(* Logix 5000 project; controller PLC_MCC1300_75F1 vendor 1 type 14 code 166 rev 32.11; software revision 32.04; part 51 of 83 *)
(* tags used below, declared in another part *)
   GP_ScadaPlate : GP_ScadaPlate;
   M310B : MAC_Conveyor;
   M310B_ALM : MAC_Conveyor_ALM;
   M310B_Data : UDT_Convoy_SL;
   M310B_HMR : MAC_Conveyor_HMR;
   M310B_SpaceConv_Utilities : SpaceConv_Utilities;
   M310Popup : MAC_Popup_ZC[2];
   M310Popup_ALM : MAC_Popup_ZC_ALM[2];
   M310Popup_HMR : MAC_Popup_ZC_HMR[2];
   M310Popup_HMW : MAC_Popup_ZC_HMW[2];
   TMP_dHalfConveyorLength : DINT;
   xAlwaysOFF : BOOL;
   xAlwaysON : BOOL;
   Z300_Conveyor : UDT_StandConv[29];
   Z300_LineTracking : UDT_LINE_TRACKING;
   Z301 : MAC_Zone_ML;
   Z401_HMI_rgtPlateScada_Internal : HMI_LiteData[5,2,7];
(* MainProgram, continued *)

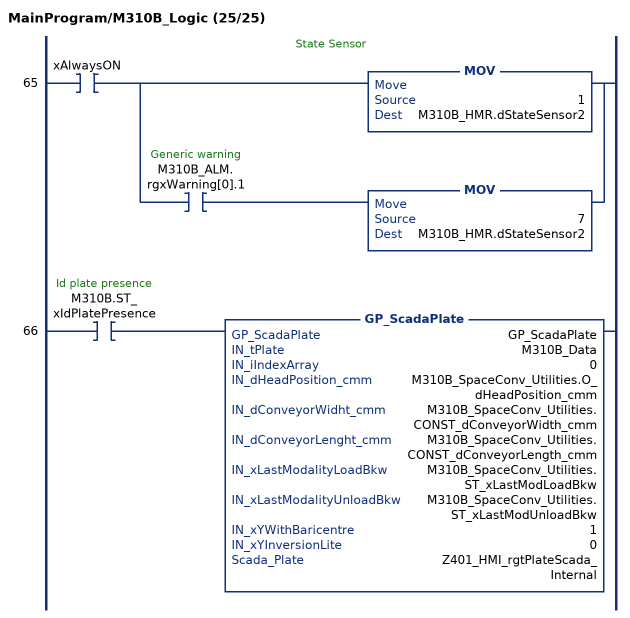
   [picture p787: MainProgram/M310B_Logic rungs 65-66]
   // State Sensor
   65: XIC(xAlwaysON)[MOV(1,M310B_HMR.dStateSensor2) ,XIC(M310B_ALM.rgxWarning[0].1) MOV(7,M310B_HMR.dStateSensor2) ];
   66: XIC(M310B.ST_xIdPlatePresence)GP_ScadaPlate(GP_ScadaPlate,M310B_Data,0,M310B_SpaceConv_Utilities.O_dHeadPosition_cmm,M310B_SpaceConv_Utilities.CONST_dConveyorWidth_cmm,M310B_SpaceConv_Utilities.CONST_dConveyorLength_cmm,M310B_SpaceConv_Utilities.ST_xLastModLoadBkw,M310B_SpaceConv_Utilities.ST_xLastModUnloadBkw,1,0,Z401_HMI_rgtPlateScada_Internal);
END_ROUTINE

ROUTINE M310Popup0_Faults   (* ladder *)
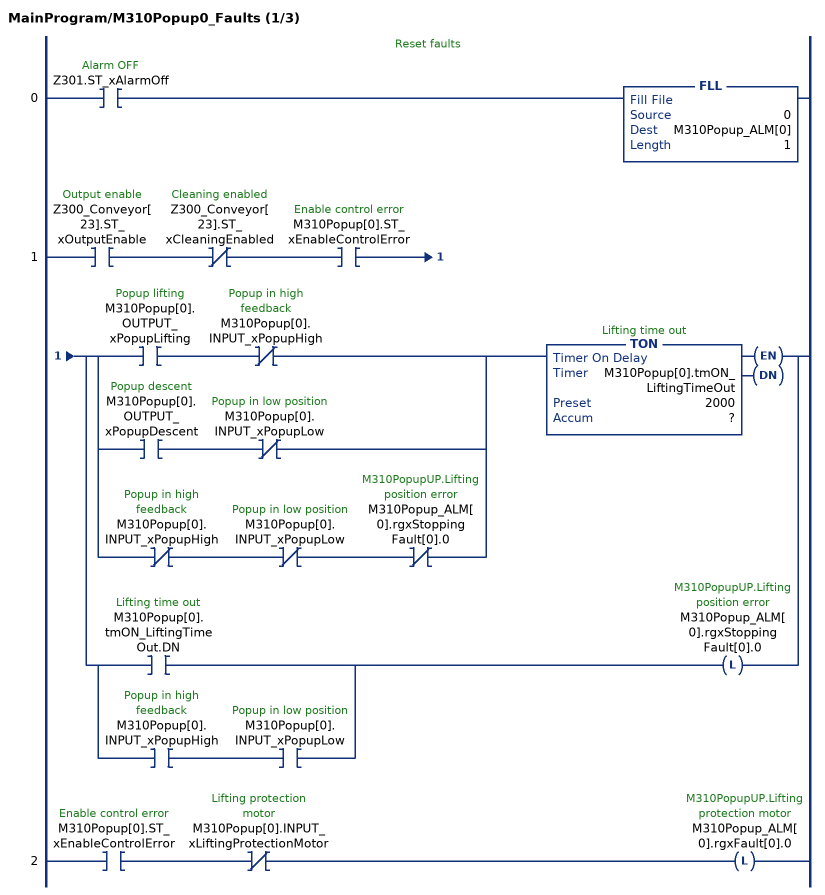
   // Reset faults
   0: XIC(Z301.ST_xAlarmOff)FLL(0,M310Popup_ALM[0],1);
   1: XIC(Z300_Conveyor[23].ST_xOutputEnable)XIO(Z300_Conveyor[23].ST_xCleaningEnabled)XIC(M310Popup[0].ST_xEnableControlError)[[XIC(M310Popup[0].OUTPUT_xPopupLifting) XIO(M310Popup[0].INPUT_xPopupHigh) ,XIC(M310Popup[0].OUTPUT_xPopupDescent) XIO(M310Popup[0].INPUT_xPopupLow) ,XIO(M310Popup[0].INPUT_xPopupHigh) XIO(M310Popup[0].INPUT_xPopupLow) XIO(M310Popup_ALM[0].rgxStoppingFault[0].0) ] TON(M310Popup[0].tmON_LiftingTimeOut,?,?) ,[XIC(M310Popup[0].tmON_LiftingTimeOut.DN) ,XIC(M310Popup[0].INPUT_xPopupHigh) XIC(M310Popup[0].INPUT_xPopupLow) ] OTL(M310Popup_ALM[0].rgxStoppingFault[0].0) ];
   2: XIC(M310Popup[0].ST_xEnableControlError)XIO(M310Popup[0].INPUT_xLiftingProtectionMotor)OTL(M310Popup_ALM[0].rgxFault[0].0);
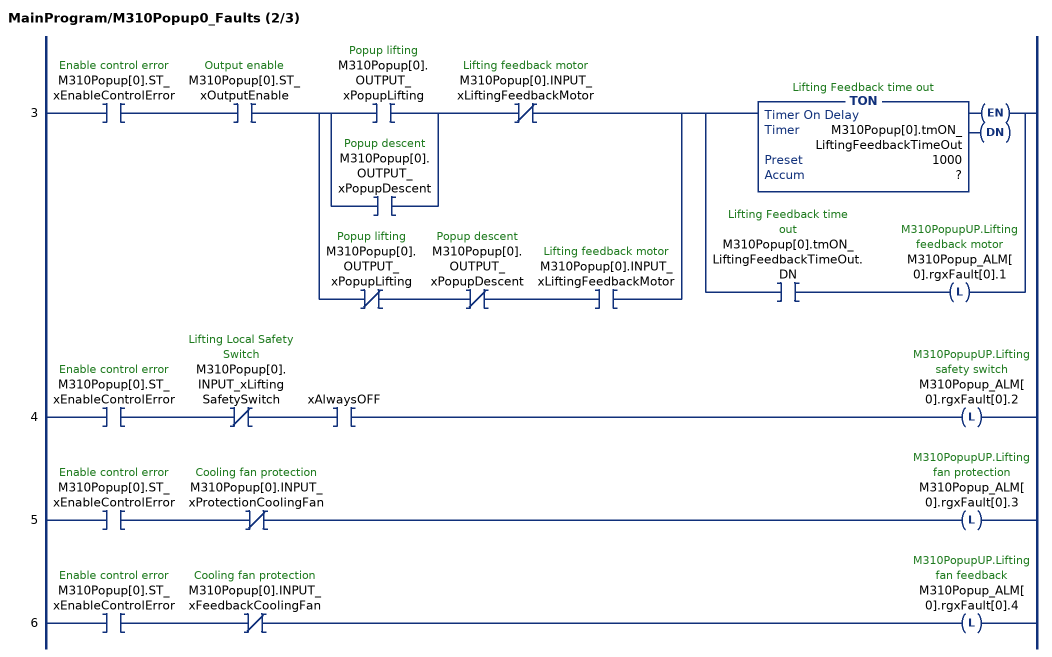
   3: XIC(M310Popup[0].ST_xEnableControlError)XIC(M310Popup[0].ST_xOutputEnable)[[XIC(M310Popup[0].OUTPUT_xPopupLifting) ,XIC(M310Popup[0].OUTPUT_xPopupDescent) ] XIO(M310Popup[0].INPUT_xLiftingFeedbackMotor) ,XIO(M310Popup[0].OUTPUT_xPopupLifting) XIO(M310Popup[0].OUTPUT_xPopupDescent) XIC(M310Popup[0].INPUT_xLiftingFeedbackMotor) ][TON(M310Popup[0].tmON_LiftingFeedbackTimeOut,?,?) ,XIC(M310Popup[0].tmON_LiftingFeedbackTimeOut.DN) OTL(M310Popup_ALM[0].rgxFault[0].1) ];
   4: XIC(M310Popup[0].ST_xEnableControlError)XIO(M310Popup[0].INPUT_xLiftingSafetySwitch)XIC(xAlwaysOFF)OTL(M310Popup_ALM[0].rgxFault[0].2);
   5: XIC(M310Popup[0].ST_xEnableControlError)XIO(M310Popup[0].INPUT_xProtectionCoolingFan)OTL(M310Popup_ALM[0].rgxFault[0].3);
   6: XIC(M310Popup[0].ST_xEnableControlError)XIO(M310Popup[0].INPUT_xFeedbackCoolingFan)OTL(M310Popup_ALM[0].rgxFault[0].4);
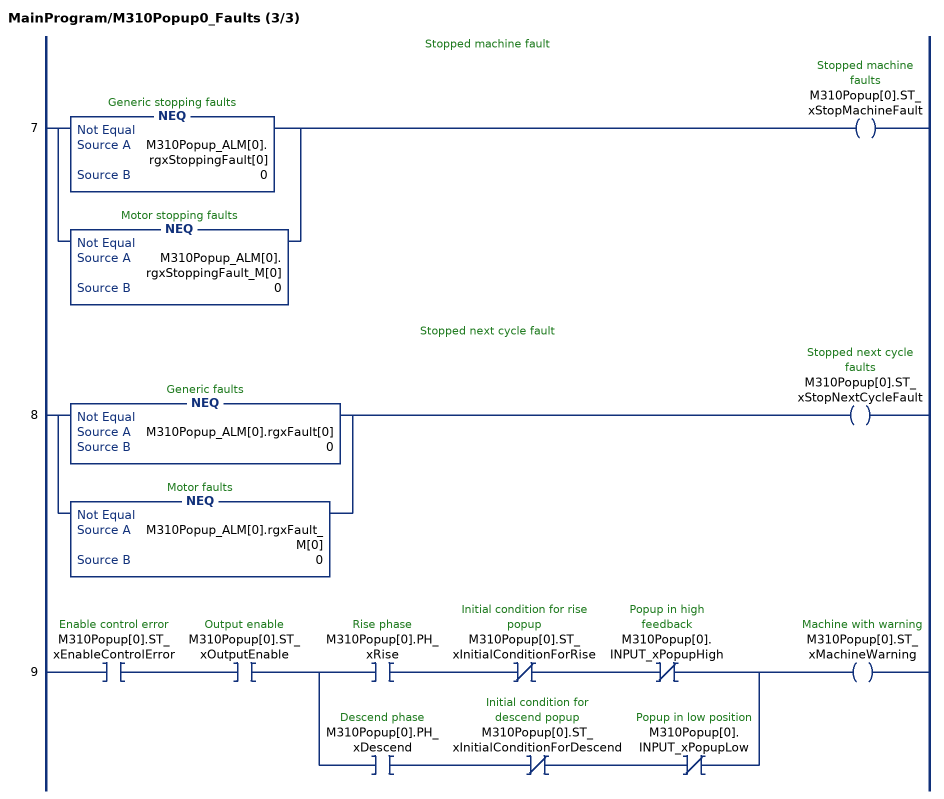
   // Stopped machine fault
   7: [NEQ(M310Popup_ALM[0].rgxStoppingFault[0],0) ,NEQ(M310Popup_ALM[0].rgxStoppingFault_M[0],0) ]OTE(M310Popup[0].ST_xStopMachineFault);
   // Stopped next cycle fault
   8: [NEQ(M310Popup_ALM[0].rgxFault[0],0) ,NEQ(M310Popup_ALM[0].rgxFault_M[0],0) ]OTE(M310Popup[0].ST_xStopNextCycleFault);
   9: XIC(M310Popup[0].ST_xEnableControlError)XIC(M310Popup[0].ST_xOutputEnable)[XIC(M310Popup[0].PH_xRise) XIO(M310Popup[0].ST_xInitialConditionForRise) XIO(M310Popup[0].INPUT_xPopupHigh) ,XIC(M310Popup[0].PH_xDescend) XIO(M310Popup[0].ST_xInitialConditionForDescend) XIO(M310Popup[0].INPUT_xPopupLow) ]OTE(M310Popup[0].ST_xMachineWarning);
END_ROUTINE

ROUTINE M310Popup0_Logic   (* ladder *)
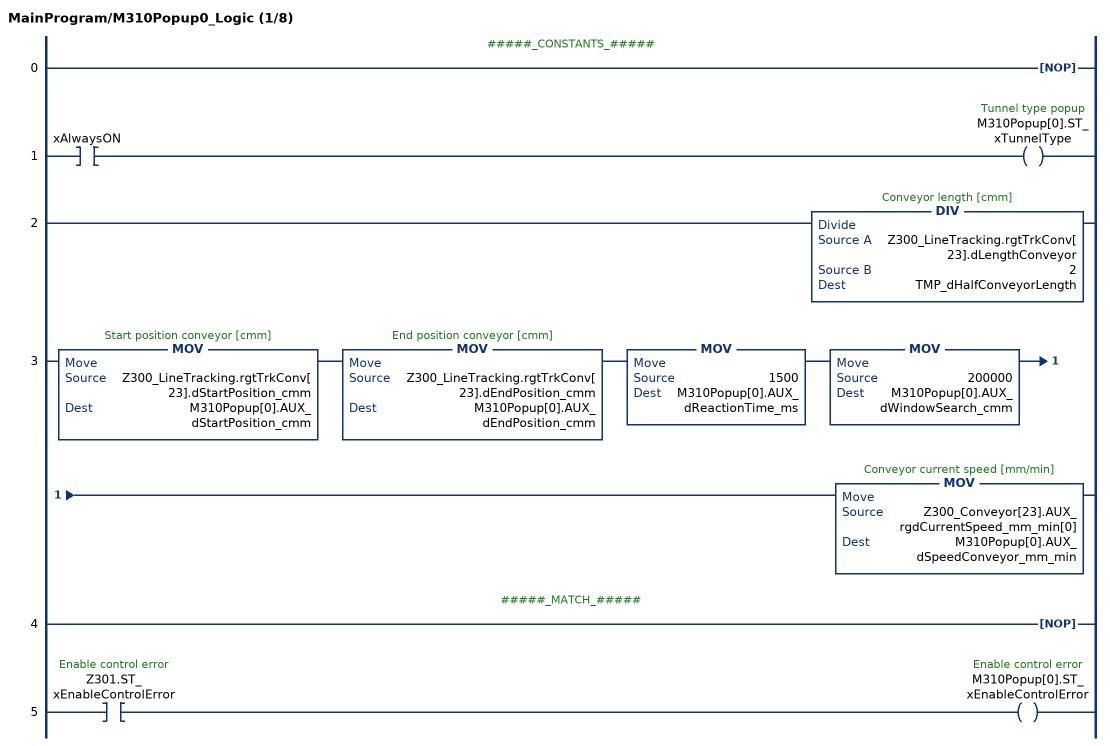
   // #####_CONSTANTS_#####
   0: NOP();
   1: XIC(xAlwaysON)OTE(M310Popup[0].ST_xTunnelType);
   2: DIV(Z300_LineTracking.rgtTrkConv[23].dLengthConveyor,2,TMP_dHalfConveyorLength);
   3: MOV(Z300_LineTracking.rgtTrkConv[23].dStartPosition_cmm,M310Popup[0].AUX_dStartPosition_cmm)MOV(Z300_LineTracking.rgtTrkConv[23].dEndPosition_cmm,M310Popup[0].AUX_dEndPosition_cmm)MOV(1500,M310Popup[0].AUX_dReactionTime_ms)MOV(200000,M310Popup[0].AUX_dWindowSearch_cmm)MOV(Z300_Conveyor[23].AUX_rgdCurrentSpeed_mm_min[0],M310Popup[0].AUX_dSpeedConveyor_mm_min);
   // #####_MATCH_#####
   4: NOP();
   5: XIC(Z301.ST_xEnableControlError)OTE(M310Popup[0].ST_xEnableControlError);
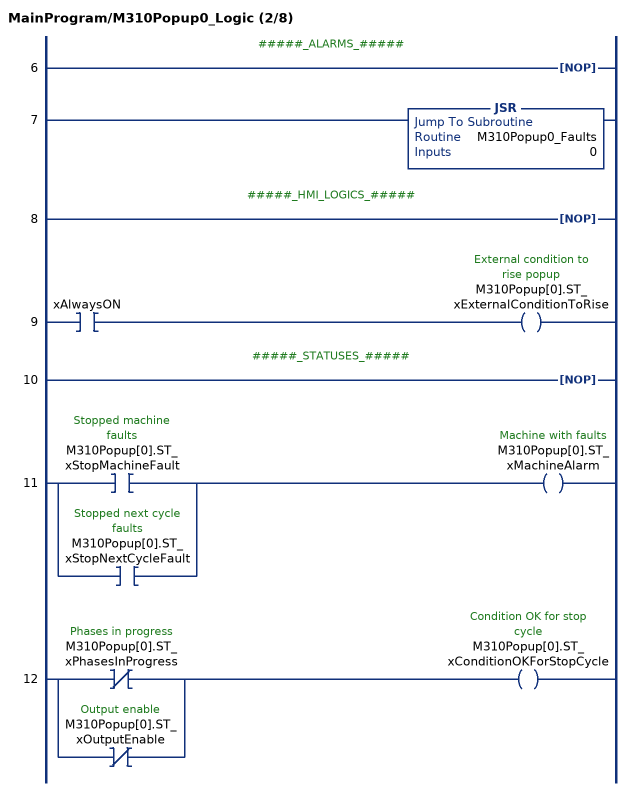
   // #####_ALARMS_#####
   6: NOP();
   7: JSR(M310Popup0_Faults,0);
   // #####_HMI_LOGICS_#####
   8: NOP();
   9: XIC(xAlwaysON)OTE(M310Popup[0].ST_xExternalConditionToRise);
   // #####_STATUSES_#####
   10: NOP();
   11: [XIC(M310Popup[0].ST_xStopMachineFault) ,XIC(M310Popup[0].ST_xStopNextCycleFault) ]OTE(M310Popup[0].ST_xMachineAlarm);
   12: [XIO(M310Popup[0].ST_xPhasesInProgress) ,XIO(M310Popup[0].ST_xOutputEnable) ]OTE(M310Popup[0].ST_xConditionOKForStopCycle);
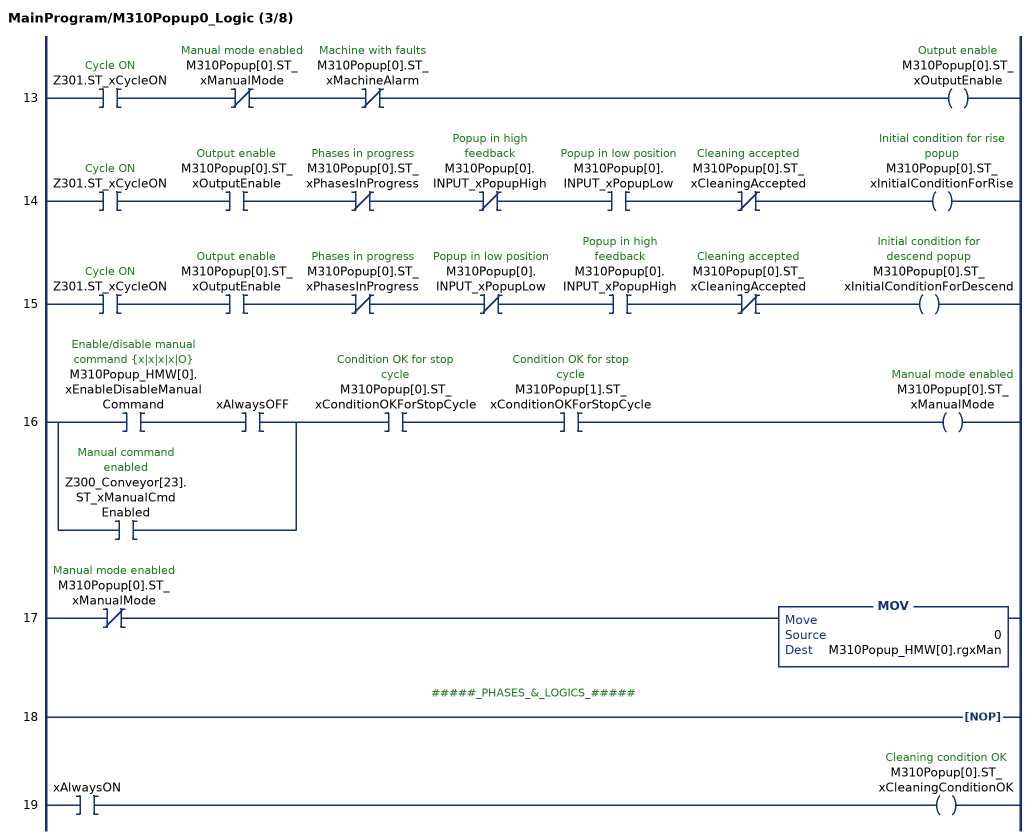
   13: XIC(Z301.ST_xCycleON)XIO(M310Popup[0].ST_xManualMode)XIO(M310Popup[0].ST_xMachineAlarm)OTE(M310Popup[0].ST_xOutputEnable);
   14: XIC(Z301.ST_xCycleON)XIC(M310Popup[0].ST_xOutputEnable)XIO(M310Popup[0].ST_xPhasesInProgress)XIO(M310Popup[0].INPUT_xPopupHigh)XIC(M310Popup[0].INPUT_xPopupLow)XIO(M310Popup[0].ST_xCleaningAccepted)OTE(M310Popup[0].ST_xInitialConditionForRise);
   15: XIC(Z301.ST_xCycleON)XIC(M310Popup[0].ST_xOutputEnable)XIO(M310Popup[0].ST_xPhasesInProgress)XIO(M310Popup[0].INPUT_xPopupLow)XIC(M310Popup[0].INPUT_xPopupHigh)XIO(M310Popup[0].ST_xCleaningAccepted)OTE(M310Popup[0].ST_xInitialConditionForDescend);
   16: [XIC(M310Popup_HMW[0].xEnableDisableManualCommand) XIC(xAlwaysOFF) ,XIC(Z300_Conveyor[23].ST_xManualCmdEnabled) ]XIC(M310Popup[0].ST_xConditionOKForStopCycle)XIC(M310Popup[1].ST_xConditionOKForStopCycle)OTE(M310Popup[0].ST_xManualMode);
   17: XIO(M310Popup[0].ST_xManualMode)MOV(0,M310Popup_HMW[0].rgxMan);
   // #####_PHASES_&_LOGICS_#####
   18: NOP();
   19: XIC(xAlwaysON)OTE(M310Popup[0].ST_xCleaningConditionOK);
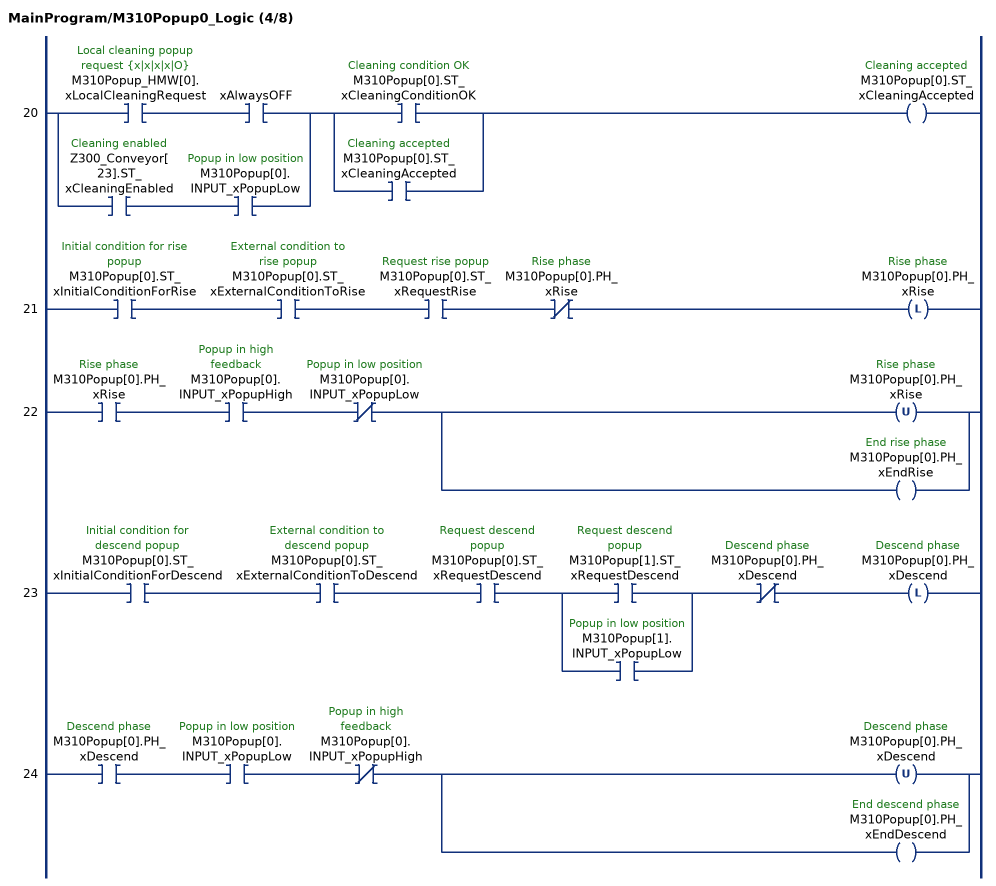
   20: [XIC(M310Popup_HMW[0].xLocalCleaningRequest) XIC(xAlwaysOFF) ,XIC(Z300_Conveyor[23].ST_xCleaningEnabled) XIC(M310Popup[0].INPUT_xPopupLow) ][XIC(M310Popup[0].ST_xCleaningConditionOK) ,XIC(M310Popup[0].ST_xCleaningAccepted) ]OTE(M310Popup[0].ST_xCleaningAccepted);
   21: XIC(M310Popup[0].ST_xInitialConditionForRise)XIC(M310Popup[0].ST_xExternalConditionToRise)XIC(M310Popup[0].ST_xRequestRise)XIO(M310Popup[0].PH_xRise)OTL(M310Popup[0].PH_xRise);
   22: XIC(M310Popup[0].PH_xRise)XIC(M310Popup[0].INPUT_xPopupHigh)XIO(M310Popup[0].INPUT_xPopupLow)[OTU(M310Popup[0].PH_xRise) ,OTE(M310Popup[0].PH_xEndRise) ];
   23: XIC(M310Popup[0].ST_xInitialConditionForDescend)XIC(M310Popup[0].ST_xExternalConditionToDescend)XIC(M310Popup[0].ST_xRequestDescend)[XIC(M310Popup[1].ST_xRequestDescend) ,XIC(M310Popup[1].INPUT_xPopupLow) ]XIO(M310Popup[0].PH_xDescend)OTL(M310Popup[0].PH_xDescend);
   24: XIC(M310Popup[0].PH_xDescend)XIC(M310Popup[0].INPUT_xPopupLow)XIO(M310Popup[0].INPUT_xPopupHigh)[OTU(M310Popup[0].PH_xDescend) ,OTE(M310Popup[0].PH_xEndDescend) ];
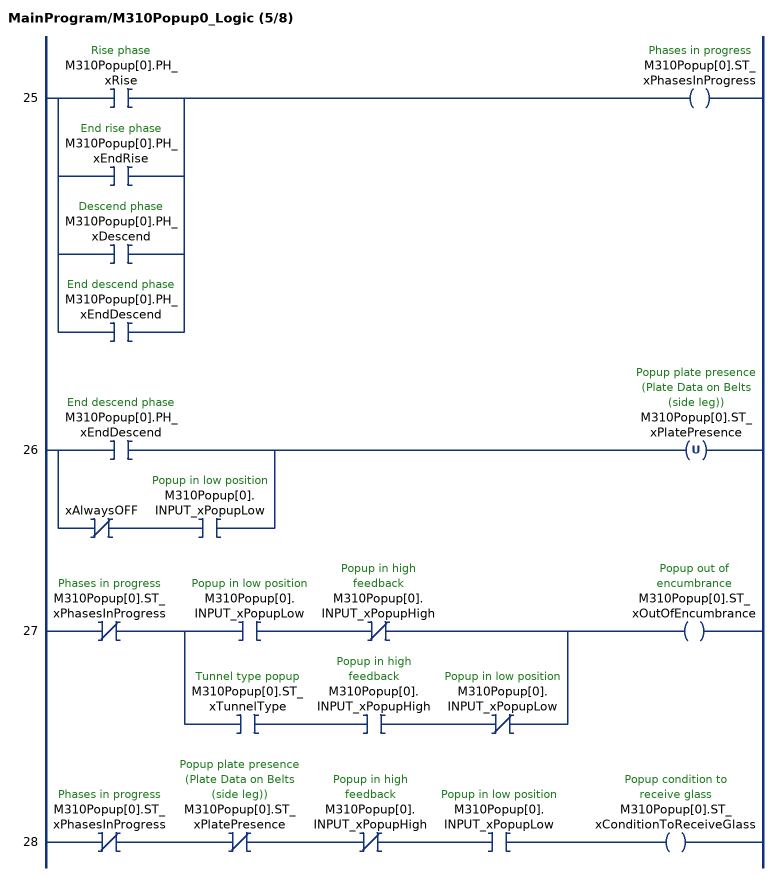
   25: [XIC(M310Popup[0].PH_xRise) ,XIC(M310Popup[0].PH_xEndRise) ,XIC(M310Popup[0].PH_xDescend) ,XIC(M310Popup[0].PH_xEndDescend) ]OTE(M310Popup[0].ST_xPhasesInProgress);
   26: [XIC(M310Popup[0].PH_xEndDescend) ,XIO(xAlwaysOFF) XIC(M310Popup[0].INPUT_xPopupLow) ]OTU(M310Popup[0].ST_xPlatePresence);
   27: XIO(M310Popup[0].ST_xPhasesInProgress)[XIC(M310Popup[0].INPUT_xPopupLow) XIO(M310Popup[0].INPUT_xPopupHigh) ,XIC(M310Popup[0].ST_xTunnelType) XIC(M310Popup[0].INPUT_xPopupHigh) XIO(M310Popup[0].INPUT_xPopupLow) ]OTE(M310Popup[0].ST_xOutOfEncumbrance);
   28: XIO(M310Popup[0].ST_xPhasesInProgress)XIO(M310Popup[0].ST_xPlatePresence)XIO(M310Popup[0].INPUT_xPopupHigh)XIC(M310Popup[0].INPUT_xPopupLow)OTE(M310Popup[0].ST_xConditionToReceiveGlass);
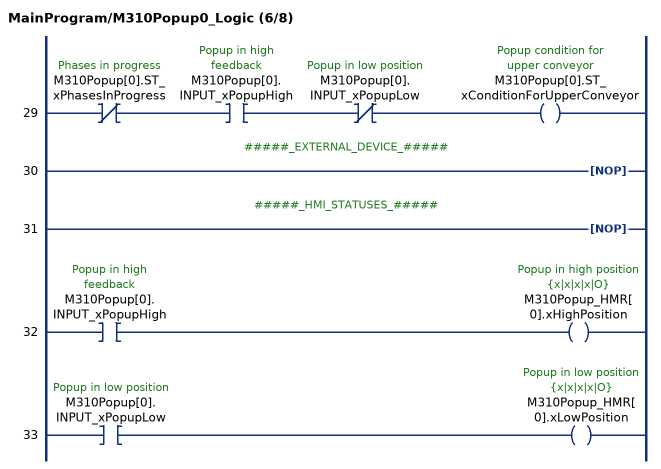
   29: XIO(M310Popup[0].ST_xPhasesInProgress)XIC(M310Popup[0].INPUT_xPopupHigh)XIO(M310Popup[0].INPUT_xPopupLow)OTE(M310Popup[0].ST_xConditionForUpperConveyor);
   // #####_EXTERNAL_DEVICE_#####
   30: NOP();
   // #####_HMI_STATUSES_#####
   31: NOP();
   32: XIC(M310Popup[0].INPUT_xPopupHigh)OTE(M310Popup_HMR[0].xHighPosition);
   33: XIC(M310Popup[0].INPUT_xPopupLow)OTE(M310Popup_HMR[0].xLowPosition);
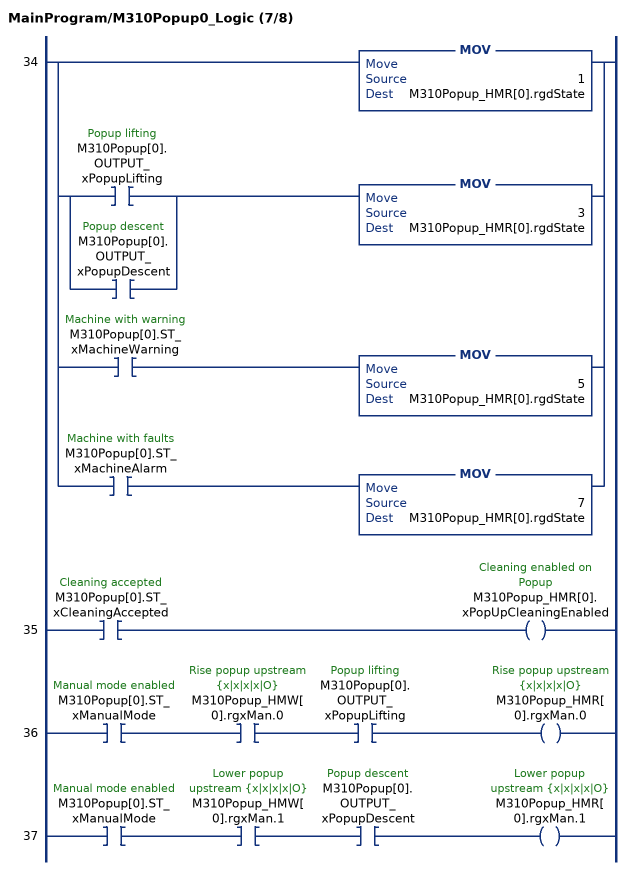
   34: [MOV(1,M310Popup_HMR[0].rgdState) ,[XIC(M310Popup[0].OUTPUT_xPopupLifting) ,XIC(M310Popup[0].OUTPUT_xPopupDescent) ] MOV(3,M310Popup_HMR[0].rgdState) ,XIC(M310Popup[0].ST_xMachineWarning) MOV(5,M310Popup_HMR[0].rgdState) ,XIC(M310Popup[0].ST_xMachineAlarm) MOV(7,M310Popup_HMR[0].rgdState) ];
   35: XIC(M310Popup[0].ST_xCleaningAccepted)OTE(M310Popup_HMR[0].xPopUpCleaningEnabled);
   36: XIC(M310Popup[0].ST_xManualMode)XIC(M310Popup_HMW[0].rgxMan.0)XIC(M310Popup[0].OUTPUT_xPopupLifting)OTE(M310Popup_HMR[0].rgxMan.0);
   37: XIC(M310Popup[0].ST_xManualMode)XIC(M310Popup_HMW[0].rgxMan.1)XIC(M310Popup[0].OUTPUT_xPopupDescent)OTE(M310Popup_HMR[0].rgxMan.1);
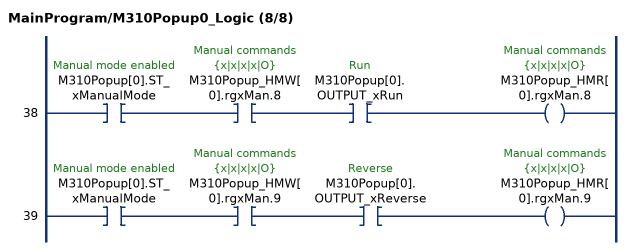
   38: XIC(M310Popup[0].ST_xManualMode)XIC(M310Popup_HMW[0].rgxMan.8)XIC(M310Popup[0].OUTPUT_xRun)OTE(M310Popup_HMR[0].rgxMan.8);
   39: XIC(M310Popup[0].ST_xManualMode)XIC(M310Popup_HMW[0].rgxMan.9)XIC(M310Popup[0].OUTPUT_xReverse)OTE(M310Popup_HMR[0].rgxMan.9);
END_ROUTINE

ROUTINE M310Popup1_Faults   (* ladder *)
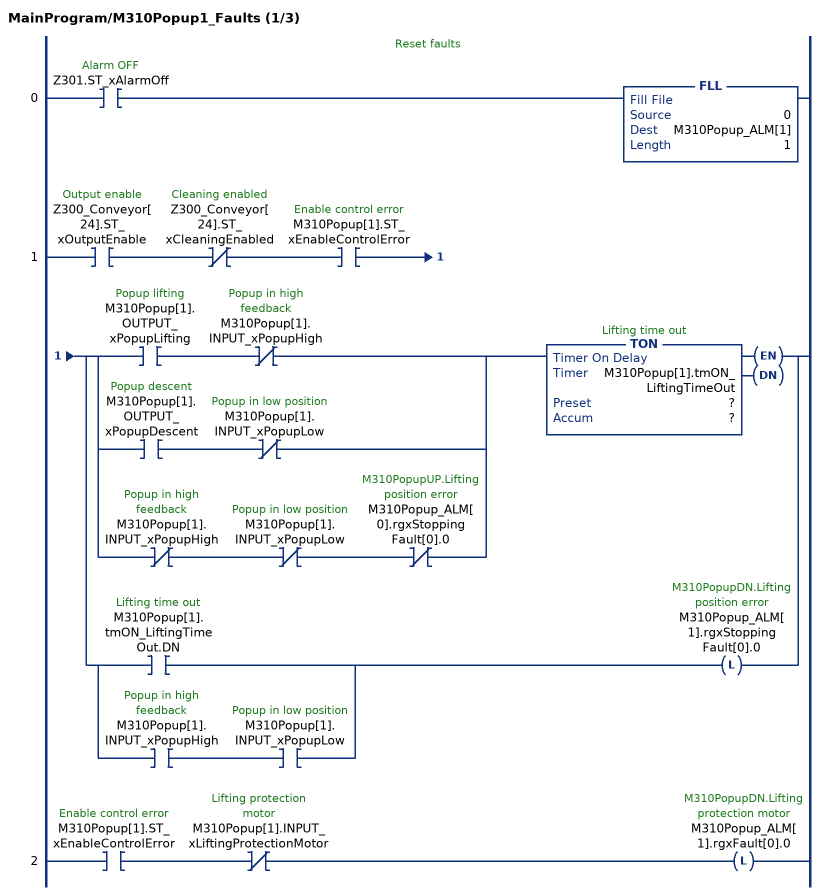
   // Reset faults
   0: XIC(Z301.ST_xAlarmOff)FLL(0,M310Popup_ALM[1],1);
   1: XIC(Z300_Conveyor[24].ST_xOutputEnable)XIO(Z300_Conveyor[24].ST_xCleaningEnabled)XIC(M310Popup[1].ST_xEnableControlError)[[XIC(M310Popup[1].OUTPUT_xPopupLifting) XIO(M310Popup[1].INPUT_xPopupHigh) ,XIC(M310Popup[1].OUTPUT_xPopupDescent) XIO(M310Popup[1].INPUT_xPopupLow) ,XIO(M310Popup[1].INPUT_xPopupHigh) XIO(M310Popup[1].INPUT_xPopupLow) XIO(M310Popup_ALM[0].rgxStoppingFault[0].0) ] TON(M310Popup[1].tmON_LiftingTimeOut,?,?) ,[XIC(M310Popup[1].tmON_LiftingTimeOut.DN) ,XIC(M310Popup[1].INPUT_xPopupHigh) XIC(M310Popup[1].INPUT_xPopupLow) ] OTL(M310Popup_ALM[1].rgxStoppingFault[0].0) ];
   2: XIC(M310Popup[1].ST_xEnableControlError)XIO(M310Popup[1].INPUT_xLiftingProtectionMotor)OTL(M310Popup_ALM[1].rgxFault[0].0);
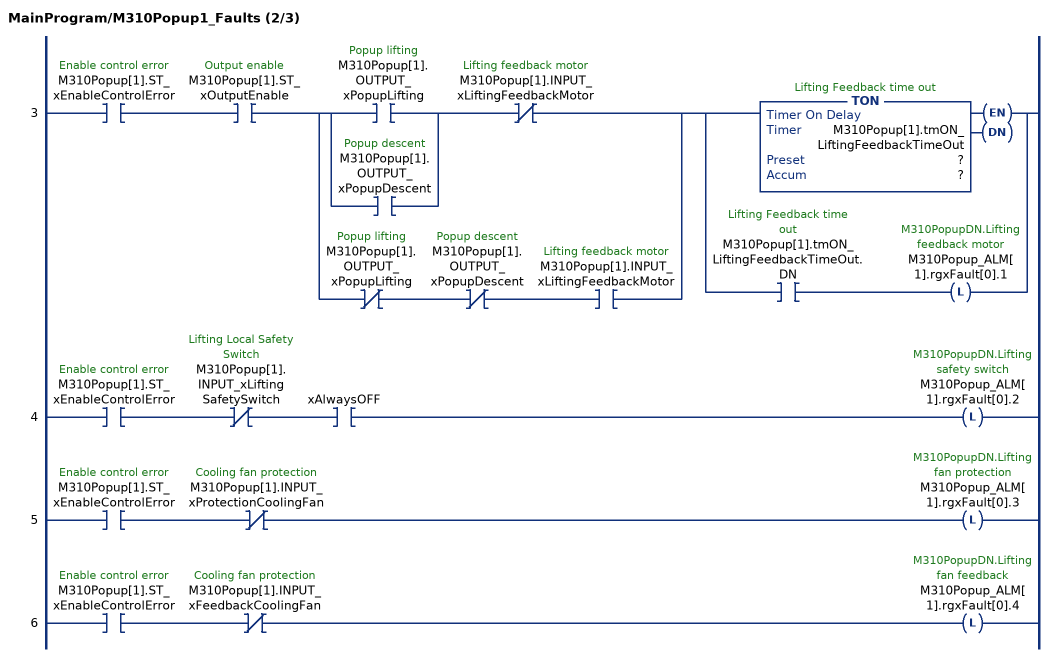
   3: XIC(M310Popup[1].ST_xEnableControlError)XIC(M310Popup[1].ST_xOutputEnable)[[XIC(M310Popup[1].OUTPUT_xPopupLifting) ,XIC(M310Popup[1].OUTPUT_xPopupDescent) ] XIO(M310Popup[1].INPUT_xLiftingFeedbackMotor) ,XIO(M310Popup[1].OUTPUT_xPopupLifting) XIO(M310Popup[1].OUTPUT_xPopupDescent) XIC(M310Popup[1].INPUT_xLiftingFeedbackMotor) ][TON(M310Popup[1].tmON_LiftingFeedbackTimeOut,?,?) ,XIC(M310Popup[1].tmON_LiftingFeedbackTimeOut.DN) OTL(M310Popup_ALM[1].rgxFault[0].1) ];
   4: XIC(M310Popup[1].ST_xEnableControlError)XIO(M310Popup[1].INPUT_xLiftingSafetySwitch)XIC(xAlwaysOFF)OTL(M310Popup_ALM[1].rgxFault[0].2);
   5: XIC(M310Popup[1].ST_xEnableControlError)XIO(M310Popup[1].INPUT_xProtectionCoolingFan)OTL(M310Popup_ALM[1].rgxFault[0].3);
   6: XIC(M310Popup[1].ST_xEnableControlError)XIO(M310Popup[1].INPUT_xFeedbackCoolingFan)OTL(M310Popup_ALM[1].rgxFault[0].4);
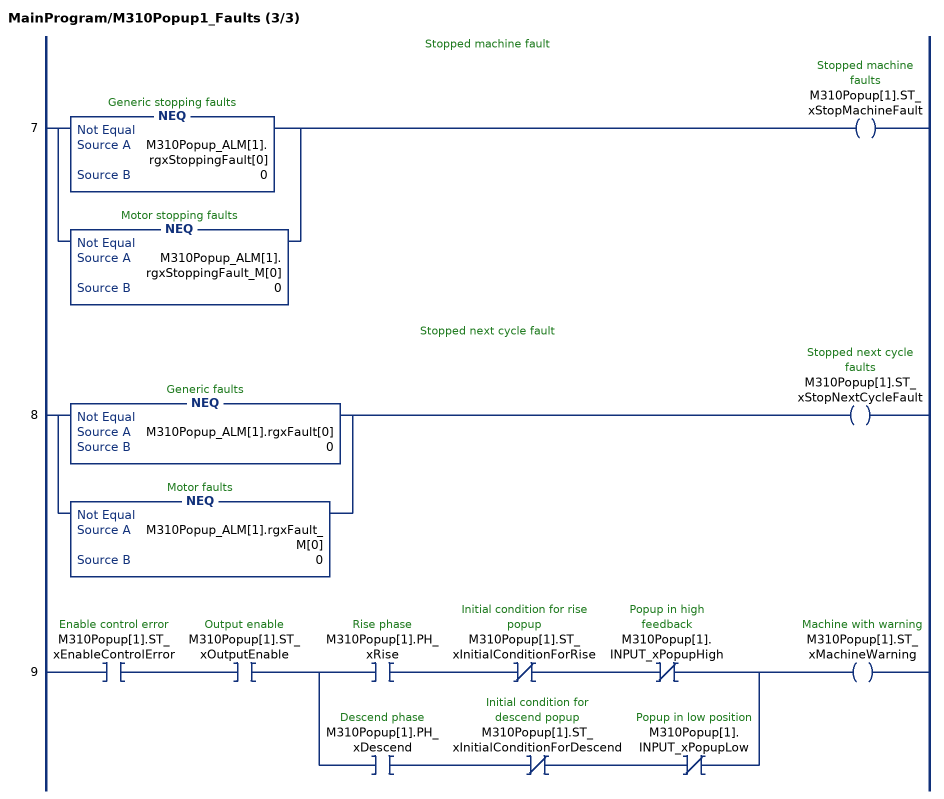
   // Stopped machine fault
   7: [NEQ(M310Popup_ALM[1].rgxStoppingFault[0],0) ,NEQ(M310Popup_ALM[1].rgxStoppingFault_M[0],0) ]OTE(M310Popup[1].ST_xStopMachineFault);
   // Stopped next cycle fault
   8: [NEQ(M310Popup_ALM[1].rgxFault[0],0) ,NEQ(M310Popup_ALM[1].rgxFault_M[0],0) ]OTE(M310Popup[1].ST_xStopNextCycleFault);
   9: XIC(M310Popup[1].ST_xEnableControlError)XIC(M310Popup[1].ST_xOutputEnable)[XIC(M310Popup[1].PH_xRise) XIO(M310Popup[1].ST_xInitialConditionForRise) XIO(M310Popup[1].INPUT_xPopupHigh) ,XIC(M310Popup[1].PH_xDescend) XIO(M310Popup[1].ST_xInitialConditionForDescend) XIO(M310Popup[1].INPUT_xPopupLow) ]OTE(M310Popup[1].ST_xMachineWarning);
END_ROUTINE

ROUTINE M310Popup1_Logic   (* ladder *)
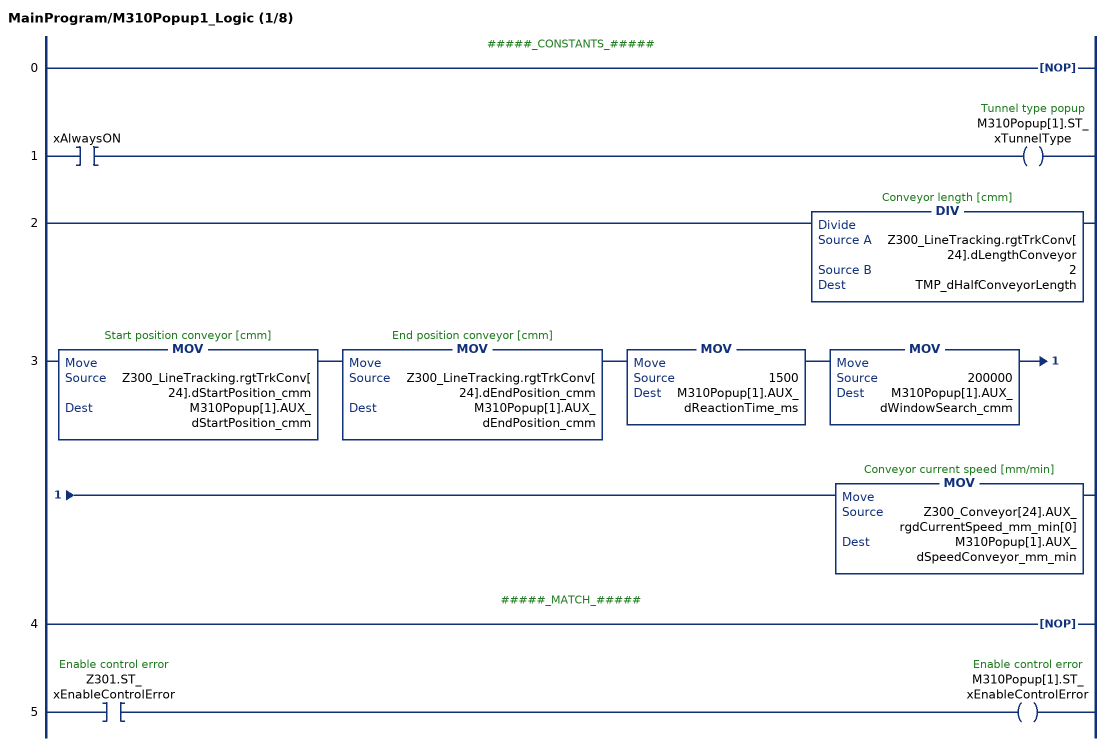
   // #####_CONSTANTS_#####
   0: NOP();
   1: XIC(xAlwaysON)OTE(M310Popup[1].ST_xTunnelType);
   2: DIV(Z300_LineTracking.rgtTrkConv[24].dLengthConveyor,2,TMP_dHalfConveyorLength);
   3: MOV(Z300_LineTracking.rgtTrkConv[24].dStartPosition_cmm,M310Popup[1].AUX_dStartPosition_cmm)MOV(Z300_LineTracking.rgtTrkConv[24].dEndPosition_cmm,M310Popup[1].AUX_dEndPosition_cmm)MOV(1500,M310Popup[1].AUX_dReactionTime_ms)MOV(200000,M310Popup[1].AUX_dWindowSearch_cmm)MOV(Z300_Conveyor[24].AUX_rgdCurrentSpeed_mm_min[0],M310Popup[1].AUX_dSpeedConveyor_mm_min);
   // #####_MATCH_#####
   4: NOP();
   5: XIC(Z301.ST_xEnableControlError)OTE(M310Popup[1].ST_xEnableControlError);
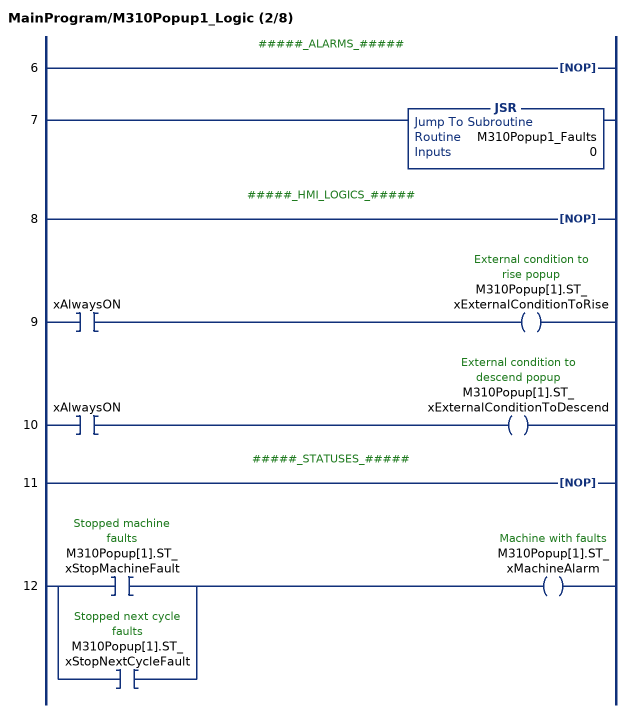
   // #####_ALARMS_#####
   6: NOP();
   7: JSR(M310Popup1_Faults,0);
   // #####_HMI_LOGICS_#####
   8: NOP();
   9: XIC(xAlwaysON)OTE(M310Popup[1].ST_xExternalConditionToRise);
   10: XIC(xAlwaysON)OTE(M310Popup[1].ST_xExternalConditionToDescend);
   // #####_STATUSES_#####
   11: NOP();
   12: [XIC(M310Popup[1].ST_xStopMachineFault) ,XIC(M310Popup[1].ST_xStopNextCycleFault) ]OTE(M310Popup[1].ST_xMachineAlarm);
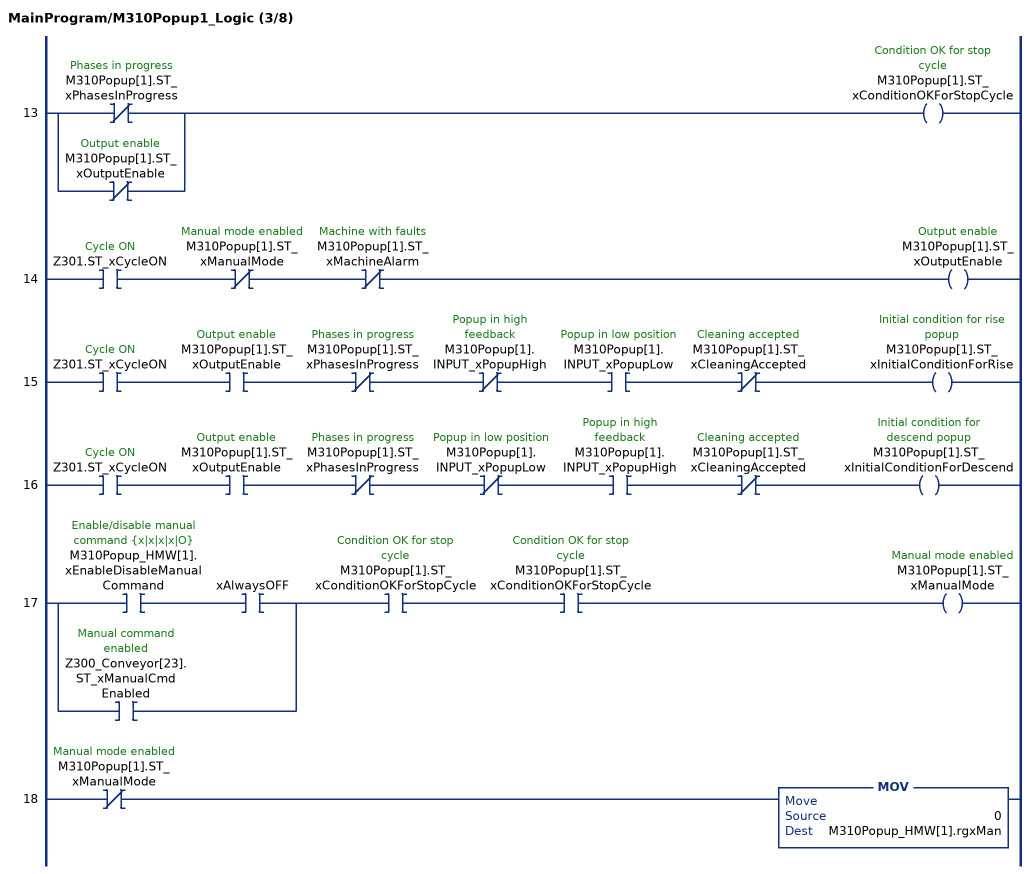
   13: [XIO(M310Popup[1].ST_xPhasesInProgress) ,XIO(M310Popup[1].ST_xOutputEnable) ]OTE(M310Popup[1].ST_xConditionOKForStopCycle);
   14: XIC(Z301.ST_xCycleON)XIO(M310Popup[1].ST_xManualMode)XIO(M310Popup[1].ST_xMachineAlarm)OTE(M310Popup[1].ST_xOutputEnable);
   15: XIC(Z301.ST_xCycleON)XIC(M310Popup[1].ST_xOutputEnable)XIO(M310Popup[1].ST_xPhasesInProgress)XIO(M310Popup[1].INPUT_xPopupHigh)XIC(M310Popup[1].INPUT_xPopupLow)XIO(M310Popup[1].ST_xCleaningAccepted)OTE(M310Popup[1].ST_xInitialConditionForRise);
   16: XIC(Z301.ST_xCycleON)XIC(M310Popup[1].ST_xOutputEnable)XIO(M310Popup[1].ST_xPhasesInProgress)XIO(M310Popup[1].INPUT_xPopupLow)XIC(M310Popup[1].INPUT_xPopupHigh)XIO(M310Popup[1].ST_xCleaningAccepted)OTE(M310Popup[1].ST_xInitialConditionForDescend);
   17: [XIC(M310Popup_HMW[1].xEnableDisableManualCommand) XIC(xAlwaysOFF) ,XIC(Z300_Conveyor[23].ST_xManualCmdEnabled) ]XIC(M310Popup[1].ST_xConditionOKForStopCycle)XIC(M310Popup[1].ST_xConditionOKForStopCycle)OTE(M310Popup[1].ST_xManualMode);
   18: XIO(M310Popup[1].ST_xManualMode)MOV(0,M310Popup_HMW[1].rgxMan);
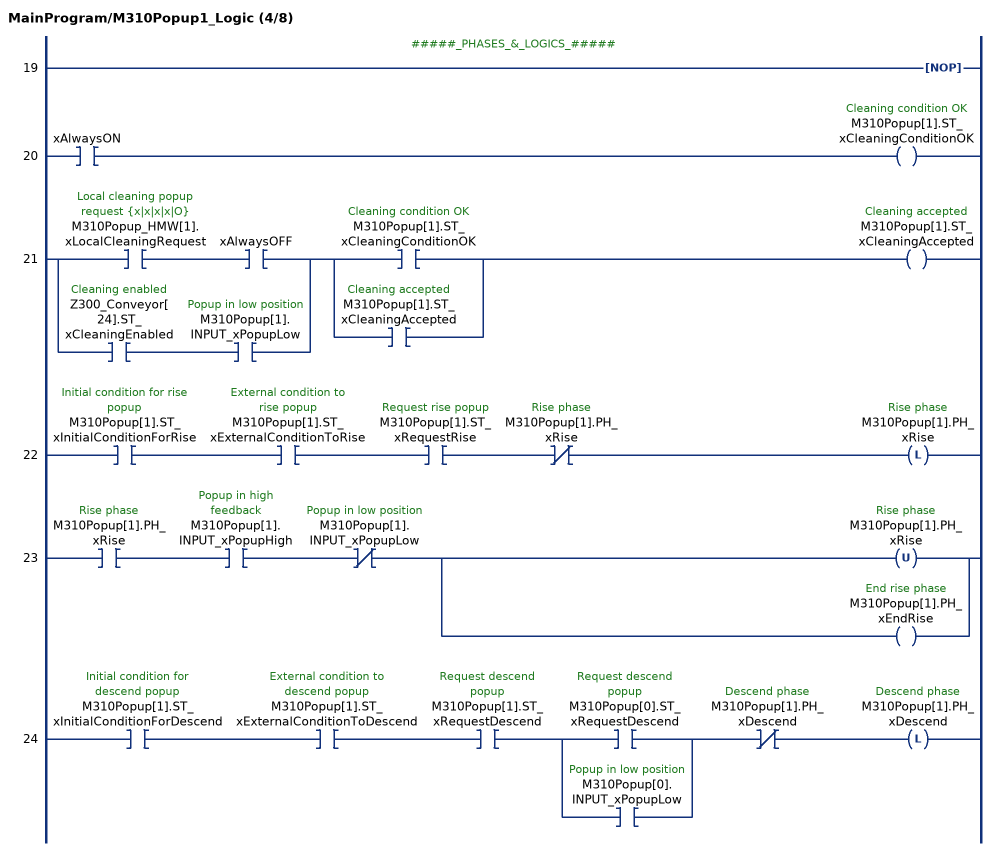
   // #####_PHASES_&_LOGICS_#####
   19: NOP();
   20: XIC(xAlwaysON)OTE(M310Popup[1].ST_xCleaningConditionOK);
   21: [XIC(M310Popup_HMW[1].xLocalCleaningRequest) XIC(xAlwaysOFF) ,XIC(Z300_Conveyor[24].ST_xCleaningEnabled) XIC(M310Popup[1].INPUT_xPopupLow) ][XIC(M310Popup[1].ST_xCleaningConditionOK) ,XIC(M310Popup[1].ST_xCleaningAccepted) ]OTE(M310Popup[1].ST_xCleaningAccepted);
   22: XIC(M310Popup[1].ST_xInitialConditionForRise)XIC(M310Popup[1].ST_xExternalConditionToRise)XIC(M310Popup[1].ST_xRequestRise)XIO(M310Popup[1].PH_xRise)OTL(M310Popup[1].PH_xRise);
   23: XIC(M310Popup[1].PH_xRise)XIC(M310Popup[1].INPUT_xPopupHigh)XIO(M310Popup[1].INPUT_xPopupLow)[OTU(M310Popup[1].PH_xRise) ,OTE(M310Popup[1].PH_xEndRise) ];
   24: XIC(M310Popup[1].ST_xInitialConditionForDescend)XIC(M310Popup[1].ST_xExternalConditionToDescend)XIC(M310Popup[1].ST_xRequestDescend)[XIC(M310Popup[0].ST_xRequestDescend) ,XIC(M310Popup[0].INPUT_xPopupLow) ]XIO(M310Popup[1].PH_xDescend)OTL(M310Popup[1].PH_xDescend);
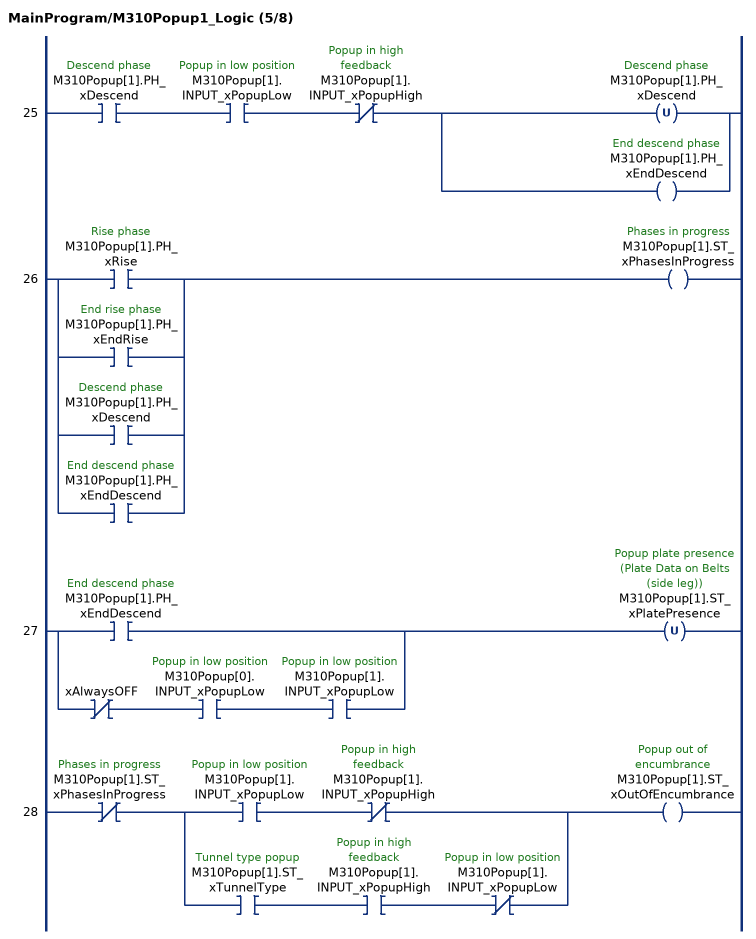
   25: XIC(M310Popup[1].PH_xDescend)XIC(M310Popup[1].INPUT_xPopupLow)XIO(M310Popup[1].INPUT_xPopupHigh)[OTU(M310Popup[1].PH_xDescend) ,OTE(M310Popup[1].PH_xEndDescend) ];
   26: [XIC(M310Popup[1].PH_xRise) ,XIC(M310Popup[1].PH_xEndRise) ,XIC(M310Popup[1].PH_xDescend) ,XIC(M310Popup[1].PH_xEndDescend) ]OTE(M310Popup[1].ST_xPhasesInProgress);
   27: [XIC(M310Popup[1].PH_xEndDescend) ,XIO(xAlwaysOFF) XIC(M310Popup[0].INPUT_xPopupLow) XIC(M310Popup[1].INPUT_xPopupLow) ]OTU(M310Popup[1].ST_xPlatePresence);
   28: XIO(M310Popup[1].ST_xPhasesInProgress)[XIC(M310Popup[1].INPUT_xPopupLow) XIO(M310Popup[1].INPUT_xPopupHigh) ,XIC(M310Popup[1].ST_xTunnelType) XIC(M310Popup[1].INPUT_xPopupHigh) XIO(M310Popup[1].INPUT_xPopupLow) ]OTE(M310Popup[1].ST_xOutOfEncumbrance);
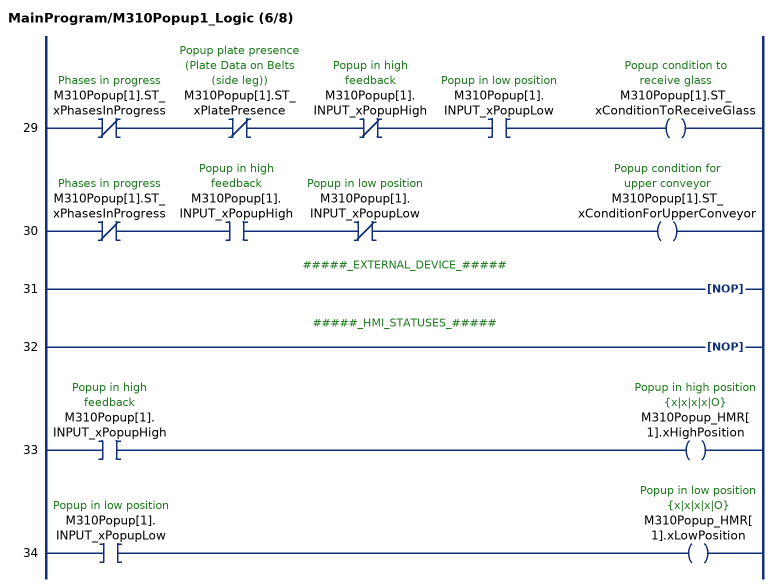
   29: XIO(M310Popup[1].ST_xPhasesInProgress)XIO(M310Popup[1].ST_xPlatePresence)XIO(M310Popup[1].INPUT_xPopupHigh)XIC(M310Popup[1].INPUT_xPopupLow)OTE(M310Popup[1].ST_xConditionToReceiveGlass);
   30: XIO(M310Popup[1].ST_xPhasesInProgress)XIC(M310Popup[1].INPUT_xPopupHigh)XIO(M310Popup[1].INPUT_xPopupLow)OTE(M310Popup[1].ST_xConditionForUpperConveyor);
   // #####_EXTERNAL_DEVICE_#####
   31: NOP();
   // #####_HMI_STATUSES_#####
   32: NOP();
   33: XIC(M310Popup[1].INPUT_xPopupHigh)OTE(M310Popup_HMR[1].xHighPosition);
   34: XIC(M310Popup[1].INPUT_xPopupLow)OTE(M310Popup_HMR[1].xLowPosition);
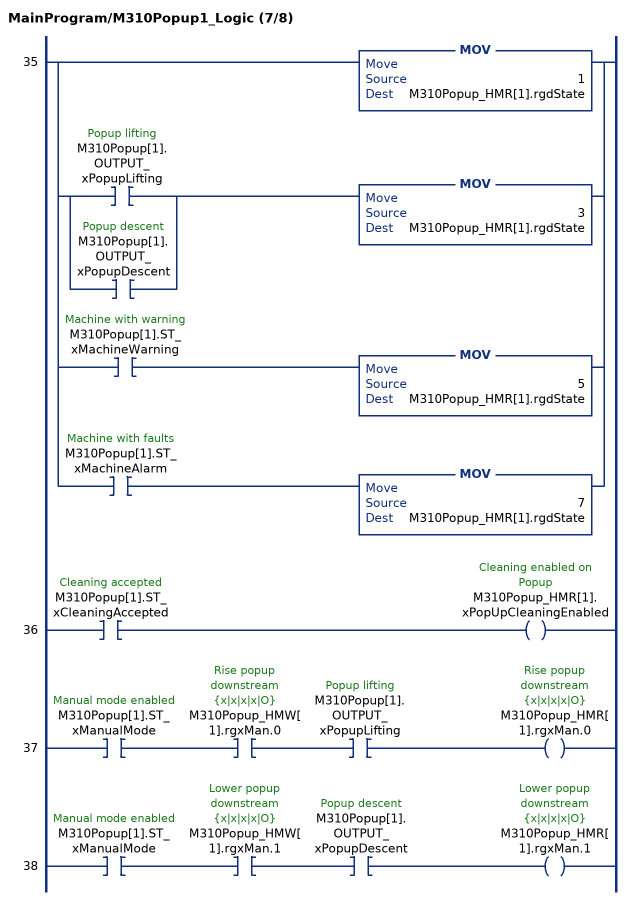
   35: [MOV(1,M310Popup_HMR[1].rgdState) ,[XIC(M310Popup[1].OUTPUT_xPopupLifting) ,XIC(M310Popup[1].OUTPUT_xPopupDescent) ] MOV(3,M310Popup_HMR[1].rgdState) ,XIC(M310Popup[1].ST_xMachineWarning) MOV(5,M310Popup_HMR[1].rgdState) ,XIC(M310Popup[1].ST_xMachineAlarm) MOV(7,M310Popup_HMR[1].rgdState) ];
   36: XIC(M310Popup[1].ST_xCleaningAccepted)OTE(M310Popup_HMR[1].xPopUpCleaningEnabled);
   37: XIC(M310Popup[1].ST_xManualMode)XIC(M310Popup_HMW[1].rgxMan.0)XIC(M310Popup[1].OUTPUT_xPopupLifting)OTE(M310Popup_HMR[1].rgxMan.0);
   38: XIC(M310Popup[1].ST_xManualMode)XIC(M310Popup_HMW[1].rgxMan.1)XIC(M310Popup[1].OUTPUT_xPopupDescent)OTE(M310Popup_HMR[1].rgxMan.1);
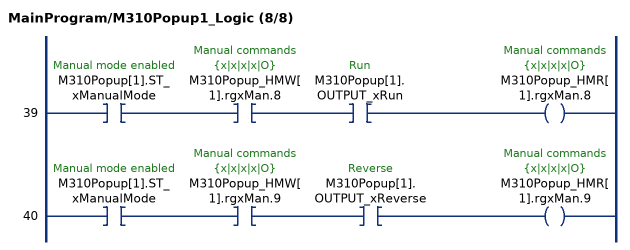
   39: XIC(M310Popup[1].ST_xManualMode)XIC(M310Popup_HMW[1].rgxMan.8)XIC(M310Popup[1].OUTPUT_xRun)OTE(M310Popup_HMR[1].rgxMan.8);
   40: XIC(M310Popup[1].ST_xManualMode)XIC(M310Popup_HMW[1].rgxMan.9)XIC(M310Popup[1].OUTPUT_xReverse)OTE(M310Popup_HMR[1].rgxMan.9);
END_ROUTINE
